REGION Network 109: ETHERNET: controllo per ripristino connessione TX
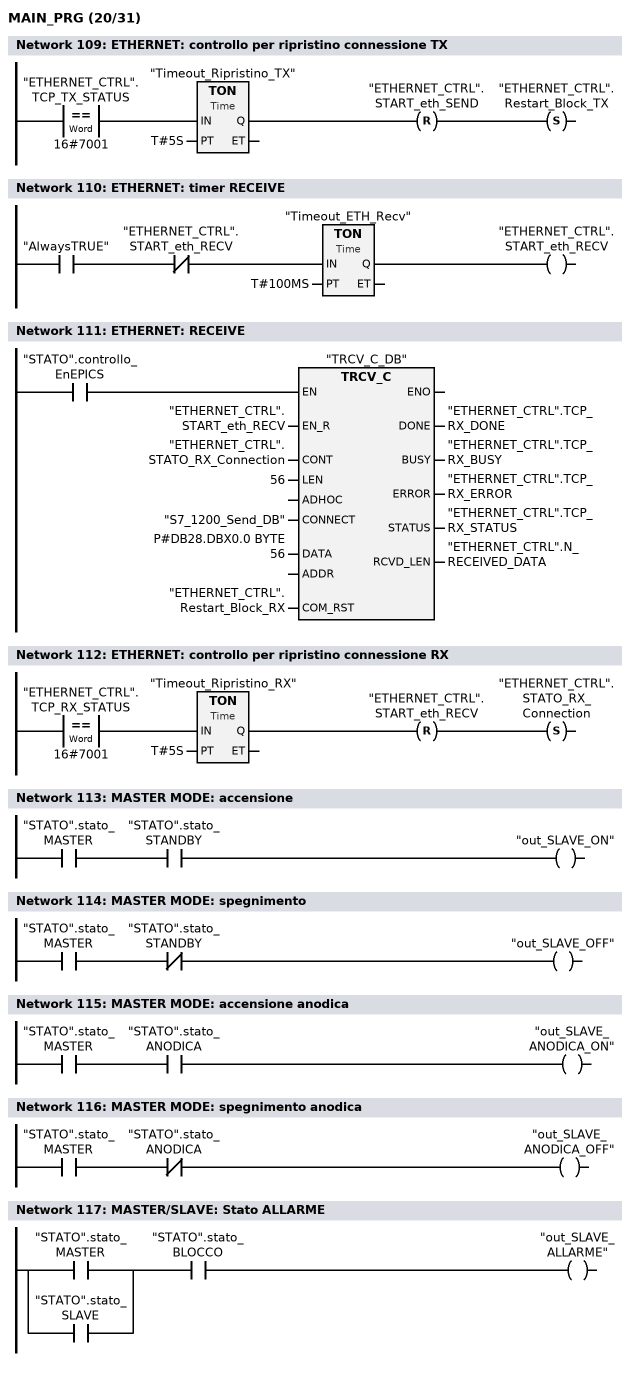
   "Timeout_Ripristino_TX".TON(IN := "ETHERNET_CTRL".TCP_TX_STATUS = 16#7001, PT := T#5S);
   IF "Timeout_Ripristino_TX".Q THEN
       "ETHERNET_CTRL".START_eth_SEND := FALSE;
       "ETHERNET_CTRL".Restart_Block_TX := TRUE;
   END_IF;
END_REGION

REGION Network 110: ETHERNET: timer RECEIVE
   "Timeout_ETH_Recv".TON(IN := "AlwaysTRUE" AND NOT "ETHERNET_CTRL".START_eth_RECV, PT := T#100MS);
   "ETHERNET_CTRL".START_eth_RECV := "Timeout_ETH_Recv".Q;
END_REGION

REGION Network 111: ETHERNET: RECEIVE
   IF "STATO".controllo_EnEPICS THEN
       "TRCV_C_DB"(EN_R := "ETHERNET_CTRL".START_eth_RECV,   // TRCV_C
                   CONT := "ETHERNET_CTRL".STATO_RX_Connection,
                   LEN := 56,
                   CONNECT := "S7_1200_Send_DB",
                   DATA := P#DB28.DBX0.0 BYTE 56,
                   COM_RST := "ETHERNET_CTRL".Restart_Block_RX,
                   DONE => "ETHERNET_CTRL".TCP_RX_DONE,
                   BUSY => "ETHERNET_CTRL".TCP_RX_BUSY,
                   ERROR => "ETHERNET_CTRL".TCP_RX_ERROR,
                   STATUS => "ETHERNET_CTRL".TCP_RX_STATUS,
                   RCVD_LEN => "ETHERNET_CTRL".N_RECEIVED_DATA);
   END_IF;
END_REGION

REGION Network 112: ETHERNET: controllo per ripristino connessione RX
   "Timeout_Ripristino_RX".TON(IN := "ETHERNET_CTRL".TCP_RX_STATUS = 16#7001, PT := T#5S);
   IF "Timeout_Ripristino_RX".Q THEN
       "ETHERNET_CTRL".START_eth_RECV := FALSE;
       "ETHERNET_CTRL".STATO_RX_Connection := TRUE;
   END_IF;
END_REGION

REGION Network 113: MASTER MODE: accensione
   RUNG wire#powerrail
      Contact( "STATO".stato_MASTER )
      Contact( "STATO".stato_STANDBY )
      Coil( "out_SLAVE_ON" )
   END_RUNG
   // the same network as SCL:
   "out_SLAVE_ON" := "STATO".stato_MASTER AND "STATO".stato_STANDBY;
END_REGION

REGION Network 114: MASTER MODE: spegnimento
   RUNG wire#powerrail
      Contact( "STATO".stato_MASTER )
      I_Contact( "STATO".stato_STANDBY )
      Coil( "out_SLAVE_OFF" )
   END_RUNG
   // the same network as SCL:
   "out_SLAVE_OFF" := "STATO".stato_MASTER AND NOT "STATO".stato_STANDBY;
END_REGION

REGION Network 115: MASTER MODE: accensione anodica
   RUNG wire#powerrail
      Contact( "STATO".stato_MASTER )
      Contact( "STATO".stato_ANODICA )
      Coil( "out_SLAVE_ANODICA_ON" )
   END_RUNG
   // the same network as SCL:
   "out_SLAVE_ANODICA_ON" := "STATO".stato_MASTER AND "STATO".stato_ANODICA;
END_REGION

REGION Network 116: MASTER MODE: spegnimento anodica
   RUNG wire#powerrail
      Contact( "STATO".stato_MASTER )
      I_Contact( "STATO".stato_ANODICA )
      Coil( "out_SLAVE_ANODICA_OFF" )
   END_RUNG
   // the same network as SCL:
   "out_SLAVE_ANODICA_OFF" := "STATO".stato_MASTER AND NOT "STATO".stato_ANODICA;
END_REGION

REGION Network 117: MASTER/SLAVE: Stato ALLARME
   RUNG wire#powerrail
      Contact( "STATO".stato_MASTER )
      wire#w1
      Contact( "STATO".stato_BLOCCO )
      Coil( "out_SLAVE_ALLARME" )
   END_RUNG
   RUNG wire#powerrail
      Contact( "STATO".stato_SLAVE )
   END_RUNG wire#w1
   // the same network as SCL:
   "out_SLAVE_ALLARME" := ("STATO".stato_MASTER OR "STATO".stato_SLAVE) AND "STATO".stato_BLOCCO;
END_REGION

REGION Network 118: MASTER/SLAVE: Stato PREALLARME
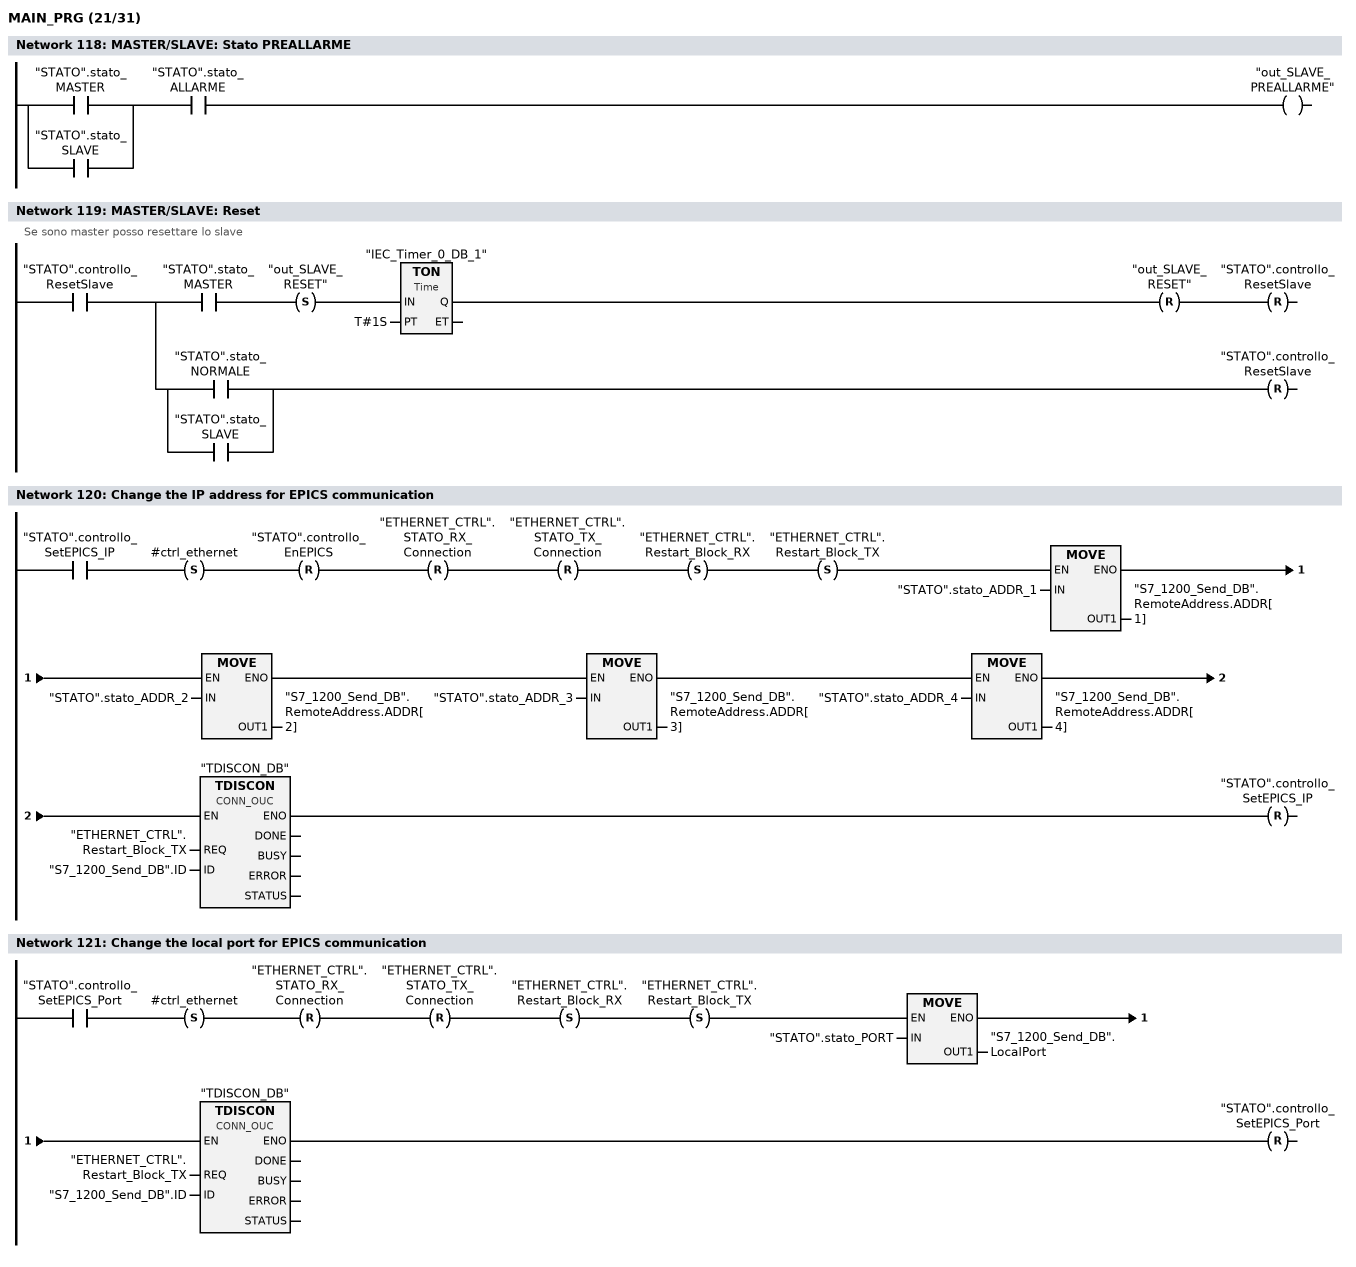
   RUNG wire#powerrail
      Contact( "STATO".stato_MASTER )
      wire#w1
      Contact( "STATO".stato_ALLARME )
      Coil( "out_SLAVE_PREALLARME" )
   END_RUNG
   RUNG wire#powerrail
      Contact( "STATO".stato_SLAVE )
   END_RUNG wire#w1
   // the same network as SCL:
   "out_SLAVE_PREALLARME" := ("STATO".stato_MASTER OR "STATO".stato_SLAVE) AND "STATO".stato_ALLARME;
END_REGION

REGION Network 119: MASTER/SLAVE: Reset
   // Se sono master posso resettare lo slave
   #_w1 := "STATO".controllo_ResetSlave AND "STATO".stato_MASTER;
   IF #_w1 THEN "out_SLAVE_RESET" := TRUE; END_IF;
   "IEC_Timer_0_DB_1".TON(IN := #_w1, PT := T#1S);
   IF "IEC_Timer_0_DB_1".Q THEN "out_SLAVE_RESET" := FALSE; END_IF;
   #_w2 := "STATO".controllo_ResetSlave;
   IF "IEC_Timer_0_DB_1".Q THEN "STATO".controllo_ResetSlave := FALSE; END_IF;
   IF #_w2 AND ("STATO".stato_NORMALE OR "STATO".stato_SLAVE) THEN
       "STATO".controllo_ResetSlave := FALSE;
   END_IF;
END_REGION

REGION Network 120: Change the IP address for EPICS communication
   // ENO of a box is taken as its EN; it also drops when the box reports an error
   IF "STATO".controllo_SetEPICS_IP THEN
       #ctrl_ethernet := TRUE;
       "STATO".controllo_EnEPICS := FALSE;
       "ETHERNET_CTRL".STATO_RX_Connection := FALSE;
       "ETHERNET_CTRL".STATO_TX_Connection := FALSE;
       "ETHERNET_CTRL".Restart_Block_RX := TRUE;
       "ETHERNET_CTRL".Restart_Block_TX := TRUE;
       "S7_1200_Send_DB".RemoteAddress.ADDR[1] := "STATO".stato_ADDR_1;
       "S7_1200_Send_DB".RemoteAddress.ADDR[2] := "STATO".stato_ADDR_2;
       "S7_1200_Send_DB".RemoteAddress.ADDR[3] := "STATO".stato_ADDR_3;
       "S7_1200_Send_DB".RemoteAddress.ADDR[4] := "STATO".stato_ADDR_4;
   END_IF;
   #_w1 := "STATO".controllo_SetEPICS_IP;
   IF #_w1 THEN
       "TDISCON_DB"(REQ := "ETHERNET_CTRL".Restart_Block_TX, ID := "S7_1200_Send_DB".ID);   // TDISCON
       "STATO".controllo_SetEPICS_IP := FALSE;
   END_IF;
END_REGION

REGION Network 121: Change the local port for EPICS communication
   // ENO of a box is taken as its EN; it also drops when the box reports an error
   IF "STATO".controllo_SetEPICS_Port THEN
       #ctrl_ethernet := TRUE;
       "ETHERNET_CTRL".STATO_RX_Connection := FALSE;
       "ETHERNET_CTRL".STATO_TX_Connection := FALSE;
       "ETHERNET_CTRL".Restart_Block_RX := TRUE;
       "ETHERNET_CTRL".Restart_Block_TX := TRUE;
       "S7_1200_Send_DB".LocalPort := "STATO".stato_PORT;
   END_IF;
   #_w1 := "STATO".controllo_SetEPICS_Port;
   IF #_w1 THEN
       "TDISCON_DB"(REQ := "ETHERNET_CTRL".Restart_Block_TX, ID := "S7_1200_Send_DB".ID);   // TDISCON
       "STATO".controllo_SetEPICS_Port := FALSE;
   END_IF;
END_REGION

REGION Network 122: Change ETHERNET parameters
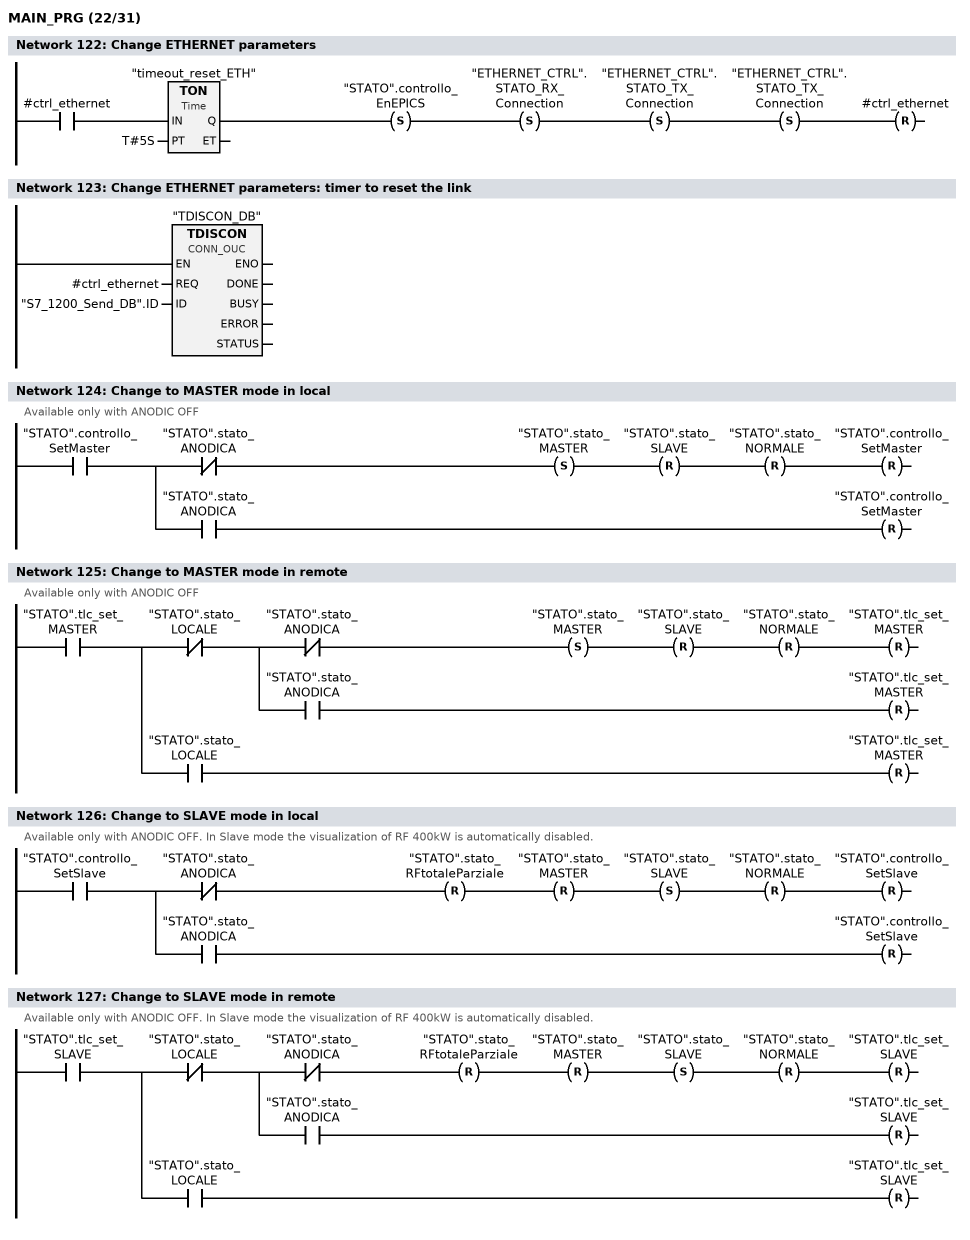
   "timeout_reset_ETH".TON(IN := #ctrl_ethernet, PT := T#5S);
   IF "timeout_reset_ETH".Q THEN
       "STATO".controllo_EnEPICS := TRUE;
       "ETHERNET_CTRL".STATO_RX_Connection := TRUE;
       "ETHERNET_CTRL".STATO_TX_Connection := TRUE;
       "ETHERNET_CTRL".STATO_TX_Connection := TRUE;
       #ctrl_ethernet := FALSE;
   END_IF;
END_REGION

REGION Network 123: Change ETHERNET parameters: timer to reset the link
   "TDISCON_DB"(REQ := #ctrl_ethernet, ID := "S7_1200_Send_DB".ID);   // TDISCON
END_REGION

REGION Network 124: Change to MASTER mode in local
   // Available only with ANODIC OFF
   RUNG wire#powerrail
      Contact( "STATO".controllo_SetMaster )
      wire#w1
      I_Contact( "STATO".stato_ANODICA )
      S_Coil( "STATO".stato_MASTER )
      R_Coil( "STATO".stato_SLAVE )
      R_Coil( "STATO".stato_NORMALE )
      R_Coil( "STATO".controllo_SetMaster )
   END_RUNG
   RUNG wire#w1
      Contact( "STATO".stato_ANODICA )
      R_Coil( "STATO".controllo_SetMaster )
   END_RUNG
   // the same network as SCL:
   IF "STATO".controllo_SetMaster AND NOT "STATO".stato_ANODICA THEN
       "STATO".stato_MASTER := TRUE;
       "STATO".stato_SLAVE := FALSE;
       "STATO".stato_NORMALE := FALSE;
   END_IF;
   #_w1 := "STATO".controllo_SetMaster;
   IF "STATO".controllo_SetMaster AND NOT "STATO".stato_ANODICA THEN
       "STATO".controllo_SetMaster := FALSE;
   END_IF;
   IF #_w1 AND "STATO".stato_ANODICA THEN "STATO".controllo_SetMaster := FALSE; END_IF;
END_REGION

REGION Network 125: Change to MASTER mode in remote
   // Available only with ANODIC OFF
   RUNG wire#powerrail
      Contact( "STATO".tlc_set_MASTER )
      wire#w1
      I_Contact( "STATO".stato_LOCALE )
      wire#w2
      I_Contact( "STATO".stato_ANODICA )
      S_Coil( "STATO".stato_MASTER )
      R_Coil( "STATO".stato_SLAVE )
      R_Coil( "STATO".stato_NORMALE )
      R_Coil( "STATO".tlc_set_MASTER )
   END_RUNG
   RUNG wire#w2
      Contact( "STATO".stato_ANODICA )
      R_Coil( "STATO".tlc_set_MASTER )
   END_RUNG
   RUNG wire#w1
      Contact( "STATO".stato_LOCALE )
      R_Coil( "STATO".tlc_set_MASTER )
   END_RUNG
   // the same network as SCL:
   #_w1 := "STATO".tlc_set_MASTER AND NOT "STATO".stato_LOCALE;
   IF #_w1 AND NOT "STATO".stato_ANODICA THEN
       "STATO".stato_MASTER := TRUE;
       "STATO".stato_SLAVE := FALSE;
       "STATO".stato_NORMALE := FALSE;
   END_IF;
   #_w2 := "STATO".tlc_set_MASTER;
   IF #_w1 AND NOT "STATO".stato_ANODICA THEN "STATO".tlc_set_MASTER := FALSE; END_IF;
   IF #_w1 AND "STATO".stato_ANODICA THEN "STATO".tlc_set_MASTER := FALSE; END_IF;
   IF #_w2 AND "STATO".stato_LOCALE THEN "STATO".tlc_set_MASTER := FALSE; END_IF;
END_REGION

REGION Network 126: Change to SLAVE mode in local
   // Available only with ANODIC OFF. In Slave mode the visualization of RF 400kW is automatically disabled.
   RUNG wire#powerrail
      Contact( "STATO".controllo_SetSlave )
      wire#w1
      I_Contact( "STATO".stato_ANODICA )
      R_Coil( "STATO".stato_RFtotaleParziale )
      R_Coil( "STATO".stato_MASTER )
      S_Coil( "STATO".stato_SLAVE )
      R_Coil( "STATO".stato_NORMALE )
      R_Coil( "STATO".controllo_SetSlave )
   END_RUNG
   RUNG wire#w1
      Contact( "STATO".stato_ANODICA )
      R_Coil( "STATO".controllo_SetSlave )
   END_RUNG
   // the same network as SCL:
   IF "STATO".controllo_SetSlave AND NOT "STATO".stato_ANODICA THEN
       "STATO".stato_RFtotaleParziale := FALSE;
       "STATO".stato_MASTER := FALSE;
       "STATO".stato_SLAVE := TRUE;
       "STATO".stato_NORMALE := FALSE;
   END_IF;
   #_w1 := "STATO".controllo_SetSlave;
   IF "STATO".controllo_SetSlave AND NOT "STATO".stato_ANODICA THEN
       "STATO".controllo_SetSlave := FALSE;
   END_IF;
   IF #_w1 AND "STATO".stato_ANODICA THEN "STATO".controllo_SetSlave := FALSE; END_IF;
END_REGION

REGION Network 127: Change to SLAVE mode in remote
   // Available only with ANODIC OFF. In Slave mode the visualization of RF 400kW is automatically disabled.
   RUNG wire#powerrail
      Contact( "STATO".tlc_set_SLAVE )
      wire#w1
      I_Contact( "STATO".stato_LOCALE )
      wire#w2
      I_Contact( "STATO".stato_ANODICA )
      R_Coil( "STATO".stato_RFtotaleParziale )
      R_Coil( "STATO".stato_MASTER )
      S_Coil( "STATO".stato_SLAVE )
      R_Coil( "STATO".stato_NORMALE )
      R_Coil( "STATO".tlc_set_SLAVE )
   END_RUNG
   RUNG wire#w2
      Contact( "STATO".stato_ANODICA )
      R_Coil( "STATO".tlc_set_SLAVE )
   END_RUNG
   RUNG wire#w1
      Contact( "STATO".stato_LOCALE )
      R_Coil( "STATO".tlc_set_SLAVE )
   END_RUNG
   // the same network as SCL:
   #_w1 := "STATO".tlc_set_SLAVE AND NOT "STATO".stato_LOCALE;
   IF #_w1 AND NOT "STATO".stato_ANODICA THEN
       "STATO".stato_RFtotaleParziale := FALSE;
       "STATO".stato_MASTER := FALSE;
       "STATO".stato_SLAVE := TRUE;
       "STATO".stato_NORMALE := FALSE;
   END_IF;
   #_w2 := "STATO".tlc_set_SLAVE;
   IF #_w1 AND NOT "STATO".stato_ANODICA THEN "STATO".tlc_set_SLAVE := FALSE; END_IF;
   IF #_w1 AND "STATO".stato_ANODICA THEN "STATO".tlc_set_SLAVE := FALSE; END_IF;
   IF #_w2 AND "STATO".stato_LOCALE THEN "STATO".tlc_set_SLAVE := FALSE; END_IF;
END_REGION

REGION Network 128: Change to NORMAL mode in local
   // Available only with ANODIC OFF. In Normal mode the visualization of RF 400kW is automatically disabled.
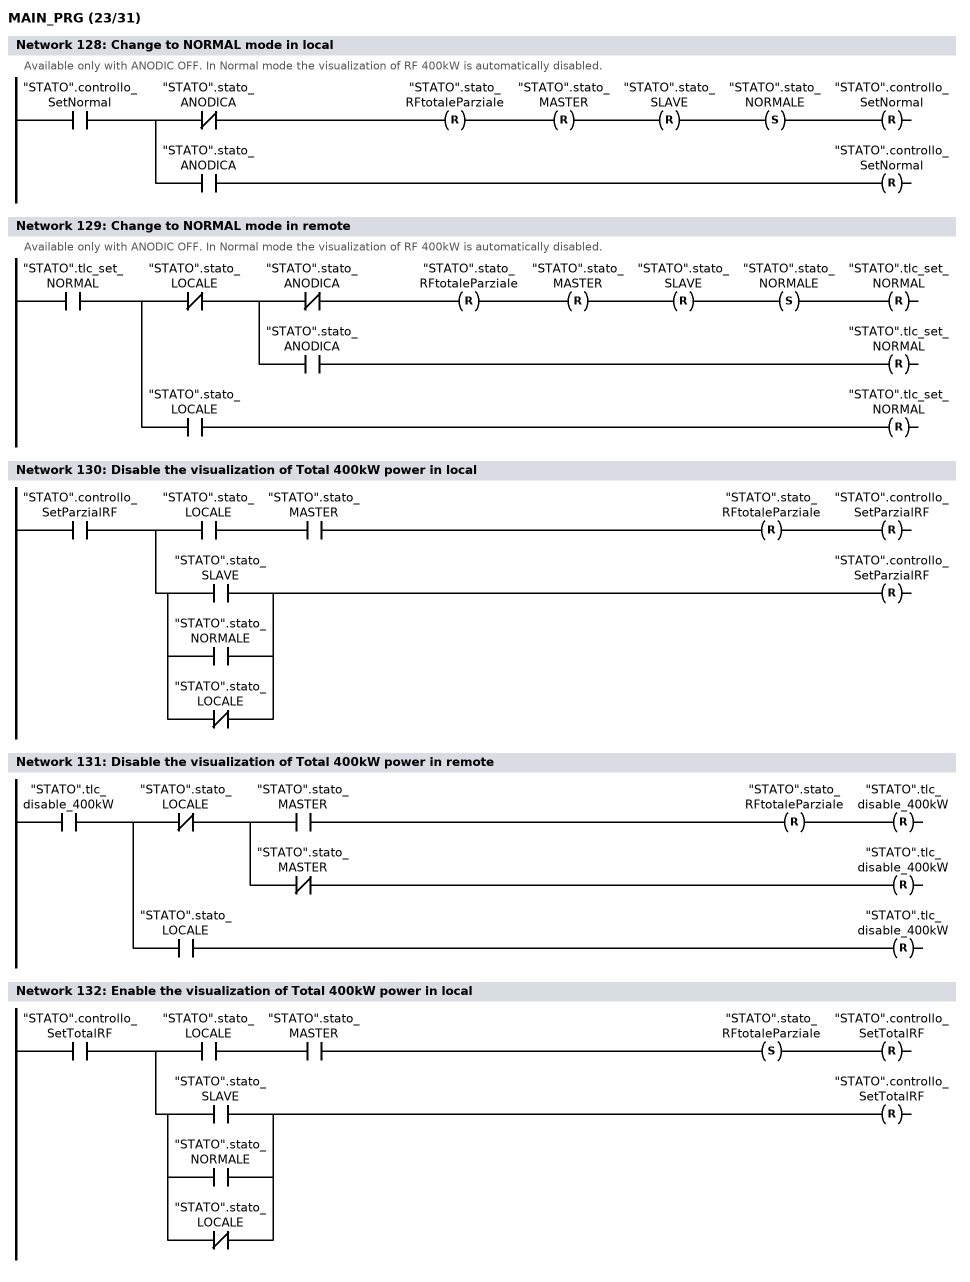
   RUNG wire#powerrail
      Contact( "STATO".controllo_SetNormal )
      wire#w1
      I_Contact( "STATO".stato_ANODICA )
      R_Coil( "STATO".stato_RFtotaleParziale )
      R_Coil( "STATO".stato_MASTER )
      R_Coil( "STATO".stato_SLAVE )
      S_Coil( "STATO".stato_NORMALE )
      R_Coil( "STATO".controllo_SetNormal )
   END_RUNG
   RUNG wire#w1
      Contact( "STATO".stato_ANODICA )
      R_Coil( "STATO".controllo_SetNormal )
   END_RUNG
   // the same network as SCL:
   IF "STATO".controllo_SetNormal AND NOT "STATO".stato_ANODICA THEN
       "STATO".stato_RFtotaleParziale := FALSE;
       "STATO".stato_MASTER := FALSE;
       "STATO".stato_SLAVE := FALSE;
       "STATO".stato_NORMALE := TRUE;
   END_IF;
   #_w1 := "STATO".controllo_SetNormal;
   IF "STATO".controllo_SetNormal AND NOT "STATO".stato_ANODICA THEN
       "STATO".controllo_SetNormal := FALSE;
   END_IF;
   IF #_w1 AND "STATO".stato_ANODICA THEN "STATO".controllo_SetNormal := FALSE; END_IF;
END_REGION

REGION Network 129: Change to NORMAL mode in remote
   // Available only with ANODIC OFF. In Normal mode the visualization of RF 400kW is automatically disabled.
   RUNG wire#powerrail
      Contact( "STATO".tlc_set_NORMAL )
      wire#w1
      I_Contact( "STATO".stato_LOCALE )
      wire#w2
      I_Contact( "STATO".stato_ANODICA )
      R_Coil( "STATO".stato_RFtotaleParziale )
      R_Coil( "STATO".stato_MASTER )
      R_Coil( "STATO".stato_SLAVE )
      S_Coil( "STATO".stato_NORMALE )
      R_Coil( "STATO".tlc_set_NORMAL )
   END_RUNG
   RUNG wire#w2
      Contact( "STATO".stato_ANODICA )
      R_Coil( "STATO".tlc_set_NORMAL )
   END_RUNG
   RUNG wire#w1
      Contact( "STATO".stato_LOCALE )
      R_Coil( "STATO".tlc_set_NORMAL )
   END_RUNG
   // the same network as SCL:
   #_w1 := "STATO".tlc_set_NORMAL AND NOT "STATO".stato_LOCALE;
   IF #_w1 AND NOT "STATO".stato_ANODICA THEN
       "STATO".stato_RFtotaleParziale := FALSE;
       "STATO".stato_MASTER := FALSE;
       "STATO".stato_SLAVE := FALSE;
       "STATO".stato_NORMALE := TRUE;
   END_IF;
   #_w2 := "STATO".tlc_set_NORMAL;
   IF #_w1 AND NOT "STATO".stato_ANODICA THEN "STATO".tlc_set_NORMAL := FALSE; END_IF;
   IF #_w1 AND "STATO".stato_ANODICA THEN "STATO".tlc_set_NORMAL := FALSE; END_IF;
   IF #_w2 AND "STATO".stato_LOCALE THEN "STATO".tlc_set_NORMAL := FALSE; END_IF;
END_REGION

REGION Network 130: Disable the visualization of Total 400kW power in local
   RUNG wire#powerrail
      Contact( "STATO".controllo_SetParzialRF )
      wire#w1
      Contact( "STATO".stato_LOCALE )
      Contact( "STATO".stato_MASTER )
      R_Coil( "STATO".stato_RFtotaleParziale )
      R_Coil( "STATO".controllo_SetParzialRF )
   END_RUNG
   RUNG wire#w1
      Contact( "STATO".stato_SLAVE )
      wire#w2
      R_Coil( "STATO".controllo_SetParzialRF )
   END_RUNG
   RUNG wire#w1
      Contact( "STATO".stato_NORMALE )
   END_RUNG wire#w2
   RUNG wire#w1
      I_Contact( "STATO".stato_LOCALE )
   END_RUNG wire#w2
   // the same network as SCL:
   IF "STATO".controllo_SetParzialRF AND "STATO".stato_LOCALE AND "STATO".stato_MASTER THEN
       "STATO".stato_RFtotaleParziale := FALSE;
   END_IF;
   #_w1 := "STATO".controllo_SetParzialRF;
   IF "STATO".controllo_SetParzialRF AND "STATO".stato_LOCALE AND "STATO".stato_MASTER THEN
       "STATO".controllo_SetParzialRF := FALSE;
   END_IF;
   IF #_w1 AND ("STATO".stato_SLAVE OR "STATO".stato_NORMALE OR NOT "STATO".stato_LOCALE) THEN
       "STATO".controllo_SetParzialRF := FALSE;
   END_IF;
END_REGION

REGION Network 131: Disable the visualization of Total 400kW power in remote
   RUNG wire#powerrail
      Contact( "STATO".tlc_disable_400kW )
      wire#w1
      I_Contact( "STATO".stato_LOCALE )
      wire#w2
      Contact( "STATO".stato_MASTER )
      R_Coil( "STATO".stato_RFtotaleParziale )
      R_Coil( "STATO".tlc_disable_400kW )
   END_RUNG
   RUNG wire#w2
      I_Contact( "STATO".stato_MASTER )
      R_Coil( "STATO".tlc_disable_400kW )
   END_RUNG
   RUNG wire#w1
      Contact( "STATO".stato_LOCALE )
      R_Coil( "STATO".tlc_disable_400kW )
   END_RUNG
   // the same network as SCL:
   #_w1 := "STATO".tlc_disable_400kW AND NOT "STATO".stato_LOCALE;
   IF #_w1 AND "STATO".stato_MASTER THEN "STATO".stato_RFtotaleParziale := FALSE; END_IF;
   #_w2 := "STATO".tlc_disable_400kW;
   IF #_w1 AND "STATO".stato_MASTER THEN "STATO".tlc_disable_400kW := FALSE; END_IF;
   IF #_w1 AND NOT "STATO".stato_MASTER THEN "STATO".tlc_disable_400kW := FALSE; END_IF;
   IF #_w2 AND "STATO".stato_LOCALE THEN "STATO".tlc_disable_400kW := FALSE; END_IF;
END_REGION

REGION Network 132: Enable the visualization of Total 400kW power in local
   RUNG wire#powerrail
      Contact( "STATO".controllo_SetTotalRF )
      wire#w1
      Contact( "STATO".stato_LOCALE )
      Contact( "STATO".stato_MASTER )
      S_Coil( "STATO".stato_RFtotaleParziale )
      R_Coil( "STATO".controllo_SetTotalRF )
   END_RUNG
   RUNG wire#w1
      Contact( "STATO".stato_SLAVE )
      wire#w2
      R_Coil( "STATO".controllo_SetTotalRF )
   END_RUNG
   RUNG wire#w1
      Contact( "STATO".stato_NORMALE )
   END_RUNG wire#w2
   RUNG wire#w1
      I_Contact( "STATO".stato_LOCALE )
   END_RUNG wire#w2
   // the same network as SCL:
   IF "STATO".controllo_SetTotalRF AND "STATO".stato_LOCALE AND "STATO".stato_MASTER THEN
       "STATO".stato_RFtotaleParziale := TRUE;
   END_IF;
   #_w1 := "STATO".controllo_SetTotalRF;
   IF "STATO".controllo_SetTotalRF AND "STATO".stato_LOCALE AND "STATO".stato_MASTER THEN
       "STATO".controllo_SetTotalRF := FALSE;
   END_IF;
   IF #_w1 AND ("STATO".stato_SLAVE OR "STATO".stato_NORMALE OR NOT "STATO".stato_LOCALE) THEN
       "STATO".controllo_SetTotalRF := FALSE;
   END_IF;
END_REGION

REGION Network 133: Enable the visualization of Total 400kW power in remote
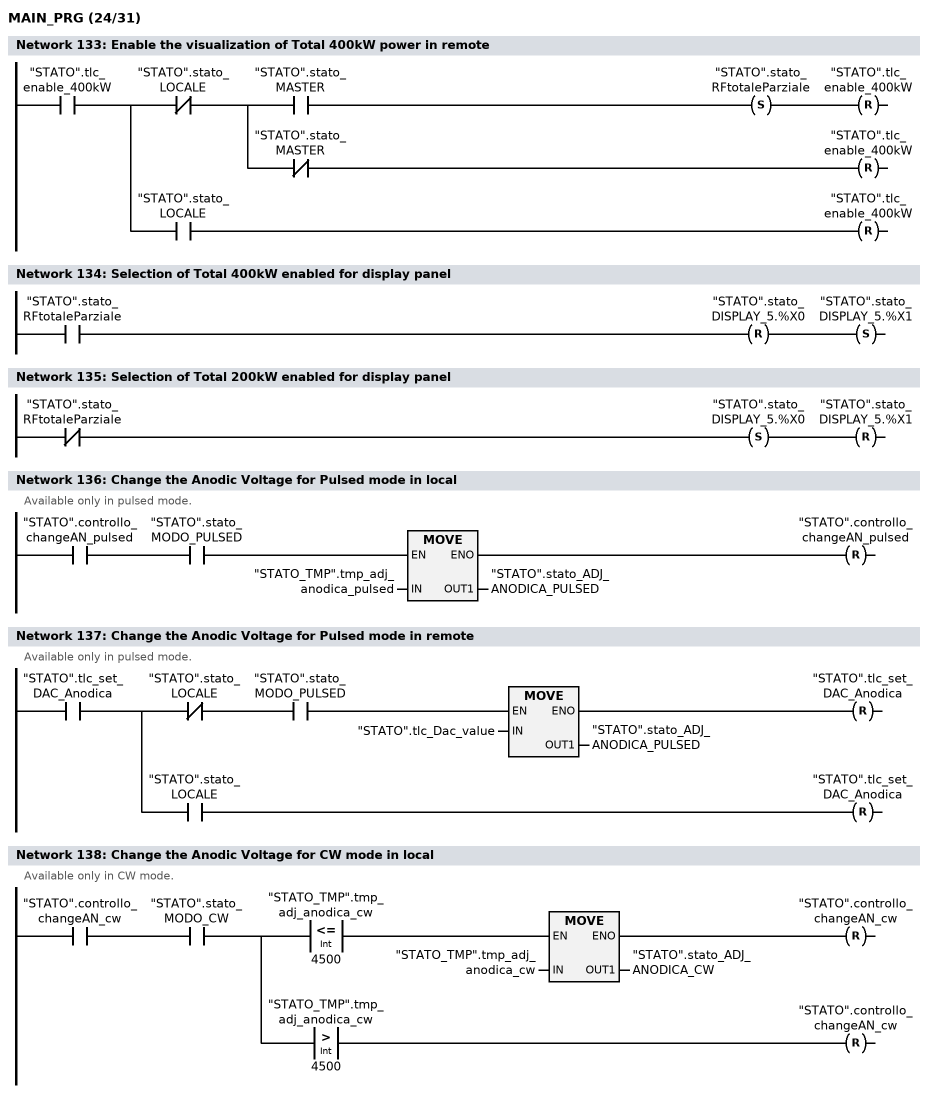
   RUNG wire#powerrail
      Contact( "STATO".tlc_enable_400kW )
      wire#w1
      I_Contact( "STATO".stato_LOCALE )
      wire#w2
      Contact( "STATO".stato_MASTER )
      S_Coil( "STATO".stato_RFtotaleParziale )
      R_Coil( "STATO".tlc_enable_400kW )
   END_RUNG
   RUNG wire#w2
      I_Contact( "STATO".stato_MASTER )
      R_Coil( "STATO".tlc_enable_400kW )
   END_RUNG
   RUNG wire#w1
      Contact( "STATO".stato_LOCALE )
      R_Coil( "STATO".tlc_enable_400kW )
   END_RUNG
   // the same network as SCL:
   #_w1 := "STATO".tlc_enable_400kW AND NOT "STATO".stato_LOCALE;
   IF #_w1 AND "STATO".stato_MASTER THEN "STATO".stato_RFtotaleParziale := TRUE; END_IF;
   #_w2 := "STATO".tlc_enable_400kW;
   IF #_w1 AND "STATO".stato_MASTER THEN "STATO".tlc_enable_400kW := FALSE; END_IF;
   IF #_w1 AND NOT "STATO".stato_MASTER THEN "STATO".tlc_enable_400kW := FALSE; END_IF;
   IF #_w2 AND "STATO".stato_LOCALE THEN "STATO".tlc_enable_400kW := FALSE; END_IF;
END_REGION

REGION Network 134: Selection of Total 400kW enabled for display panel
   RUNG wire#powerrail
      Contact( "STATO".stato_RFtotaleParziale )
      R_Coil( "STATO".stato_DISPLAY_5.%X0 )
      S_Coil( "STATO".stato_DISPLAY_5.%X1 )
   END_RUNG
   // the same network as SCL:
   IF "STATO".stato_RFtotaleParziale THEN
       "STATO".stato_DISPLAY_5.%X0 := FALSE;
       "STATO".stato_DISPLAY_5.%X1 := TRUE;
   END_IF;
END_REGION

REGION Network 135: Selection of Total 200kW enabled for display panel
   RUNG wire#powerrail
      I_Contact( "STATO".stato_RFtotaleParziale )
      S_Coil( "STATO".stato_DISPLAY_5.%X0 )
      R_Coil( "STATO".stato_DISPLAY_5.%X1 )
   END_RUNG
   // the same network as SCL:
   IF NOT "STATO".stato_RFtotaleParziale THEN
       "STATO".stato_DISPLAY_5.%X0 := TRUE;
       "STATO".stato_DISPLAY_5.%X1 := FALSE;
   END_IF;
END_REGION

REGION Network 136: Change the Anodic Voltage for Pulsed mode in local
   // Available only in pulsed mode.
   RUNG wire#powerrail
      Contact( "STATO".controllo_changeAN_pulsed )
      Contact( "STATO".stato_MODO_PULSED )
      Move(in := "STATO_TMP".tmp_adj_anodica_pulsed, out1 => "STATO".stato_ADJ_ANODICA_PULSED)
      R_Coil( "STATO".controllo_changeAN_pulsed )
   END_RUNG
   // the same network as SCL:
   IF "STATO".controllo_changeAN_pulsed AND "STATO".stato_MODO_PULSED THEN
       "STATO".stato_ADJ_ANODICA_PULSED := "STATO_TMP".tmp_adj_anodica_pulsed;
       "STATO".controllo_changeAN_pulsed := FALSE;
   END_IF;
END_REGION

REGION Network 137: Change the Anodic Voltage for Pulsed mode in remote
   // Available only in pulsed mode.
   RUNG wire#powerrail
      Contact( "STATO".tlc_set_DAC_Anodica )
      wire#w1
      I_Contact( "STATO".stato_LOCALE )
      Contact( "STATO".stato_MODO_PULSED )
      Move(in := "STATO".tlc_Dac_value, out1 => "STATO".stato_ADJ_ANODICA_PULSED)
      R_Coil( "STATO".tlc_set_DAC_Anodica )
   END_RUNG
   RUNG wire#w1
      Contact( "STATO".stato_LOCALE )
      R_Coil( "STATO".tlc_set_DAC_Anodica )
   END_RUNG
   // the same network as SCL:
   IF "STATO".tlc_set_DAC_Anodica AND NOT "STATO".stato_LOCALE AND "STATO".stato_MODO_PULSED THEN
       "STATO".stato_ADJ_ANODICA_PULSED := "STATO".tlc_Dac_value;
   END_IF;
   #_w1 := "STATO".tlc_set_DAC_Anodica;
   IF "STATO".tlc_set_DAC_Anodica AND NOT "STATO".stato_LOCALE AND "STATO".stato_MODO_PULSED THEN
       "STATO".tlc_set_DAC_Anodica := FALSE;
   END_IF;
   IF #_w1 AND "STATO".stato_LOCALE THEN "STATO".tlc_set_DAC_Anodica := FALSE; END_IF;
END_REGION

REGION Network 138: Change the Anodic Voltage for CW mode in local
   // Available only in CW mode.
   RUNG wire#powerrail
      Contact( "STATO".controllo_changeAN_cw )
      Contact( "STATO".stato_MODO_CW )
      wire#w1
      { S7_Templates := "SrcType := Int" } LE_Contact(in1 := "STATO_TMP".tmp_adj_anodica_cw, in2 := 4500)
      Move(in := "STATO_TMP".tmp_adj_anodica_cw, out1 => "STATO".stato_ADJ_ANODICA_CW)
      R_Coil( "STATO".controllo_changeAN_cw )
   END_RUNG
   RUNG wire#w1
      { S7_Templates := "SrcType := Int" } GT_Contact(in1 := "STATO_TMP".tmp_adj_anodica_cw, in2 := 4500)
      R_Coil( "STATO".controllo_changeAN_cw )
   END_RUNG
   // the same network as SCL:
   #_w1 := "STATO".controllo_changeAN_cw AND "STATO".stato_MODO_CW;
   IF #_w1 AND ("STATO_TMP".tmp_adj_anodica_cw <= 4500) THEN
       "STATO".stato_ADJ_ANODICA_CW := "STATO_TMP".tmp_adj_anodica_cw;
       "STATO".controllo_changeAN_cw := FALSE;
   END_IF;
   IF #_w1 AND ("STATO_TMP".tmp_adj_anodica_cw > 4500) THEN "STATO".controllo_changeAN_cw := FALSE; END_IF;
END_REGION

REGION Network 139: Change the Anodic Voltage for CW mode in remote
   // Available only in CW mode.
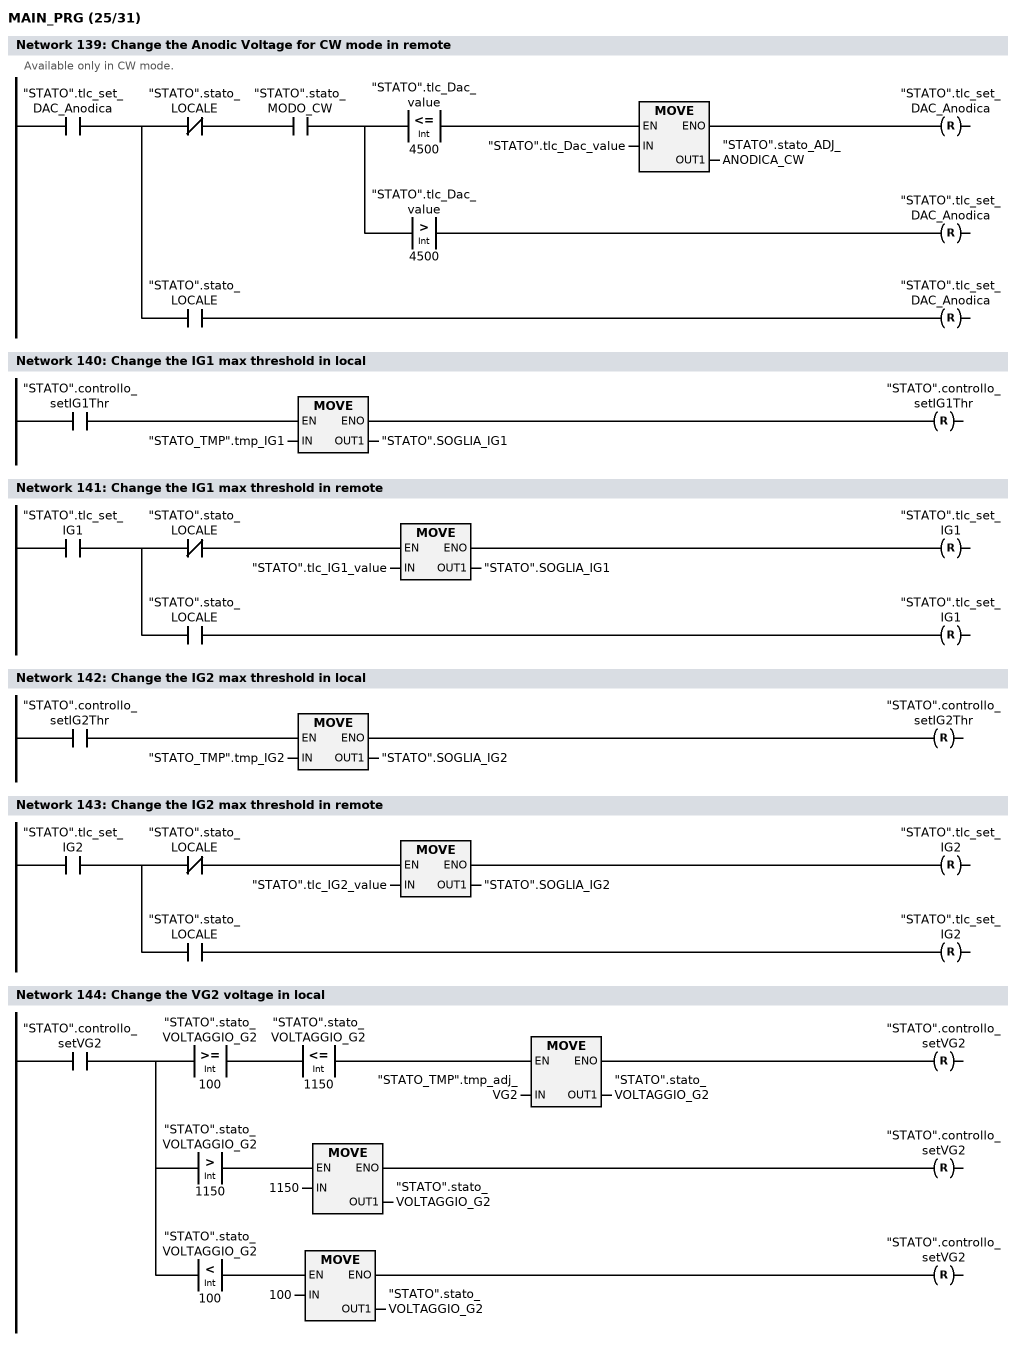
   RUNG wire#powerrail
      Contact( "STATO".tlc_set_DAC_Anodica )
      wire#w1
      I_Contact( "STATO".stato_LOCALE )
      Contact( "STATO".stato_MODO_CW )
      wire#w2
      { S7_Templates := "SrcType := Int" } LE_Contact(in1 := "STATO".tlc_Dac_value, in2 := 4500)
      Move(in := "STATO".tlc_Dac_value, out1 => "STATO".stato_ADJ_ANODICA_CW)
      R_Coil( "STATO".tlc_set_DAC_Anodica )
   END_RUNG
   RUNG wire#w2
      { S7_Templates := "SrcType := Int" } GT_Contact(in1 := "STATO".tlc_Dac_value, in2 := 4500)
      R_Coil( "STATO".tlc_set_DAC_Anodica )
   END_RUNG
   RUNG wire#w1
      Contact( "STATO".stato_LOCALE )
      R_Coil( "STATO".tlc_set_DAC_Anodica )
   END_RUNG
   // the same network as SCL:
   #_w1 := "STATO".tlc_set_DAC_Anodica AND NOT "STATO".stato_LOCALE AND "STATO".stato_MODO_CW;
   IF #_w1 AND ("STATO".tlc_Dac_value <= 4500) THEN
       "STATO".stato_ADJ_ANODICA_CW := "STATO".tlc_Dac_value;
   END_IF;
   #_w2 := "STATO".tlc_set_DAC_Anodica;
   IF #_w1 AND ("STATO".tlc_Dac_value <= 4500) THEN "STATO".tlc_set_DAC_Anodica := FALSE; END_IF;
   IF #_w1 AND ("STATO".tlc_Dac_value > 4500) THEN "STATO".tlc_set_DAC_Anodica := FALSE; END_IF;
   IF #_w2 AND "STATO".stato_LOCALE THEN "STATO".tlc_set_DAC_Anodica := FALSE; END_IF;
END_REGION

REGION Network 140: Change the IG1 max threshold in local
   RUNG wire#powerrail
      Contact( "STATO".controllo_setIG1Thr )
      Move(in := "STATO_TMP".tmp_IG1, out1 => "STATO".SOGLIA_IG1)
      R_Coil( "STATO".controllo_setIG1Thr )
   END_RUNG
   // the same network as SCL:
   IF "STATO".controllo_setIG1Thr THEN
       "STATO".SOGLIA_IG1 := "STATO_TMP".tmp_IG1;
       "STATO".controllo_setIG1Thr := FALSE;
   END_IF;
END_REGION

REGION Network 141: Change the IG1 max threshold in remote
   RUNG wire#powerrail
      Contact( "STATO".tlc_set_IG1 )
      wire#w1
      I_Contact( "STATO".stato_LOCALE )
      Move(in := "STATO".tlc_IG1_value, out1 => "STATO".SOGLIA_IG1)
      R_Coil( "STATO".tlc_set_IG1 )
   END_RUNG
   RUNG wire#w1
      Contact( "STATO".stato_LOCALE )
      R_Coil( "STATO".tlc_set_IG1 )
   END_RUNG
   // the same network as SCL:
   IF "STATO".tlc_set_IG1 AND NOT "STATO".stato_LOCALE THEN
       "STATO".SOGLIA_IG1 := "STATO".tlc_IG1_value;
   END_IF;
   #_w1 := "STATO".tlc_set_IG1;
   IF "STATO".tlc_set_IG1 AND NOT "STATO".stato_LOCALE THEN "STATO".tlc_set_IG1 := FALSE; END_IF;
   IF #_w1 AND "STATO".stato_LOCALE THEN "STATO".tlc_set_IG1 := FALSE; END_IF;
END_REGION

REGION Network 142: Change the IG2 max threshold in local
   RUNG wire#powerrail
      Contact( "STATO".controllo_setIG2Thr )
      Move(in := "STATO_TMP".tmp_IG2, out1 => "STATO".SOGLIA_IG2)
      R_Coil( "STATO".controllo_setIG2Thr )
   END_RUNG
   // the same network as SCL:
   IF "STATO".controllo_setIG2Thr THEN
       "STATO".SOGLIA_IG2 := "STATO_TMP".tmp_IG2;
       "STATO".controllo_setIG2Thr := FALSE;
   END_IF;
END_REGION

REGION Network 143: Change the IG2 max threshold in remote
   RUNG wire#powerrail
      Contact( "STATO".tlc_set_IG2 )
      wire#w1
      I_Contact( "STATO".stato_LOCALE )
      Move(in := "STATO".tlc_IG2_value, out1 => "STATO".SOGLIA_IG2)
      R_Coil( "STATO".tlc_set_IG2 )
   END_RUNG
   RUNG wire#w1
      Contact( "STATO".stato_LOCALE )
      R_Coil( "STATO".tlc_set_IG2 )
   END_RUNG
   // the same network as SCL:
   IF "STATO".tlc_set_IG2 AND NOT "STATO".stato_LOCALE THEN
       "STATO".SOGLIA_IG2 := "STATO".tlc_IG2_value;
   END_IF;
   #_w1 := "STATO".tlc_set_IG2;
   IF "STATO".tlc_set_IG2 AND NOT "STATO".stato_LOCALE THEN "STATO".tlc_set_IG2 := FALSE; END_IF;
   IF #_w1 AND "STATO".stato_LOCALE THEN "STATO".tlc_set_IG2 := FALSE; END_IF;
END_REGION
